(* Logix 5000 project; controller MV vendor 1 type 14 code 217 rev 31.11; software revision 31.00 *) (continued)
        [2].5   // Channel 1 extend button available
        [32].5   // CH1 run return flow check timer
        [26]   // CH1 no.of tank to be cleaned
        [31].0   // CH1 scavenge initialised
        [31].1   // CH1 prerinse initialised
        [32].4   // CH1 run return pump flag
        [34]   // CH1 command processor current step
        [38]   // CH1 pointer to DT service data file
        [11]   // CH1 route no.
        [33].2   // CH1 detergent tank high level probe covered
        [35]   // CH1 restart step
   MC_N100_20_alarm : ALARM_DIGITAL;
   MC_N100_20_Alarm_Ready : BOOL;
   MC_N100_20_Delayed_Timer2 : TIMER := (PRE := 1000);
   MC_N100_20_Fault_Returned : STRING;
   MC_N100_20_SQL_Done : DINT := -1;
   MC_N100_23_alarm : ALARM_DIGITAL;
   MC_N100_23_Alarm_Ready : BOOL;
   MC_N100_23_Delayed_Timer2 : TIMER := (PRE := 1000);
   MC_N100_23_Event_Returned : STRING := 'CH1_R1 feedbacks have failed.';
   MC_N100_23_Fault_Returned : STRING;
   MC_N100_23_SQL_Done : DINT := -1;
   MC_N100_29_0_Storagebit : BOOL;
   MC_N100_29_1_Storagebit : BOOL;
   MC_N100_29_2_Storagebit : BOOL;
   MC_N100_29_3_Storagebit : BOOL;
   MC_N100_29_4_Storagebit : BOOL;
   MC_N101 : INT[255];   // CH1 PC>PLC Channel 1 PC to PLC
        [0]   // CH1 PC button selected
        [0].2   // Stop channel 1 CIP selected
        [0].5   // Extend Channel 1 CIP selected
        [0].6   // Channel 1 end extend selected
        [0].15   // CH1 startup cancelled
        [0].7   // Channel 1 skip selected
        [0].4   // Abort channel 1 CIP selected
        [0].3   // Continue channel 1 CIP selected
        [0].1   // Start CH1 selected
        [0].0   // Initiate CH1 startup
   MC_N102 : INT[255] := ([1] := 1, [2] := 70, [3] := 1, [4] := 900, [5] := 1, [6] := 300, [10] := 2000, [11] := 90, [12] := 120, [13] := 7, [14] := 1, [15] := 6, [16] := 17, [17] := 1017, [19] := 11068, [21] := -1, [22] := -32768, [23] := -32768, [24] := -32768, [25] := -32768, [26] := -32768, [27] := -32768, [28] := -32768, [29] := -32768, [30] := -32768, [31] := -32768);   // CH1 PROG Channel 1 CIP progra m
        [1]   // CH1 no.prerinse cycles
        [10]   // CH1 CIP program flowrate setpoint (??/??)
        [14]   // CH1 CIP program detergent tank to use (1-2)
        [13].1   // CH1 recover rinse water flag
        [13].2   // CH1 use recovered water flag
        [0]   // CH1 scavenge time
        [15]   // CH1 CIP program route no.(1-6)
        [9]   // CH1 CIP program pressure setpoint (PSI)
        [16]   // CH1 CIP program program no.(1-47)
        [13].0   // CH1 Is Line Clean flag
        [21]   // CH1 CIP program vessel no.
        [4]   // CH1 detergent cycle time
        [6]   // CH1 postrinse cycle time
        [2]   // CH1 prerinse cycle time
        [3]   // CH1 no.detergent cycles
        [5]   // CH1 no.postrinse cycles
   MC_N103 : INT[255] := ([1] := 1, [2] := 2, [3] := 3, [4] := 4, [5] := 5, [6] := 6, [7] := 7, [8] := 8, [9] := 9, [10] := 10, [11] := 11, [12] := 12, [13] := 13, [14] := 14, [15] := 15, [16] := 16, [17] := 17, [18] := 18, [19] := 19, [20] := 64, [21] := 9999, [22] := 9999, [23] := 9999, [24] := 62, [25] := 99, [26] := -32768, [27] := 9999, [28] := 9999, [29] := 9999, [30] := 9999, [31] := -32768);   // CH1 ITEMS Chwd.nos.of items to be checked for Chan nel 1
        [0]   // CH1/R1 checkword no.
        [1]   // CH1/R2 checkword no.
        [2]   // CH1/R3 checkword no.
        [3]   // CH1/R4 checkword no.
        [4]   // CH1/R5 checkword no.
        [5]   // CH1/R6 checkword no.
        [12]   // CH1/DRAIN checkword no.
        [13]   // CH1/RR checkword no.
        [6]   // CH1/R1R checkword no.
        [7]   // CH1/R2R checkword no.
        [8]   // CH1/R3R checkword no.
        [9]   // CH1/R4R checkword no.
        [10]   // CH1/R5R checkword no.
        [11]   // CH1/R6R checkword no.
        [14]   // CH1/DR1 checkword no.
        [15]   // CH1/DR2 checkword no.
        [16]   // CH1/DT1 checkword no.
        [17]   // CH1/DT2 checkword no.
        [18]   // CH1/PR1 checkword no.
        [19]   // CH1/LF1 checkword no.
        [20]   // P1 checkword no.
   MC_N104 : INT[255] := ([0] := 6, [1] := 1017, [3] := 11068, [5] := 3, [6] := 14, [9] := 1);   // CH1 REPORT Channel 1 CIP report file
        [0].3   // CH1 final detergent strength save required
        [9]   // CH1 report detergent tank used (1 or 2)
        [0].0   // CH1 PLC -> PC save CIP report flag
        [0].1   // CH1 report save starting detergent strength flag
        [0].2   // CH1 report save final detergent strength flag
        [0]   // CH1 report flags
   MC_N108 : INT[255] := ([0] := 20, [1] := 8, [2] := 20, [3] := 4, [4] := 1);   // CH1 VDATA Channel 1 CIP progra m validation data
        [3]   // CH1 program validation loops this scan
        [4].0   // CH1 program validation complete flag
        [2]   // CH1 program validation loop counter
        [1]   // CH1 program validation max.loops per scan
        [4].1   // CH1 CIP program invalid flag
        [0]   // CH1 program validation CIP program size
        [4]   // CH1 program validation flags
   MC_N112 : INT[255] := ([0] := 1, [1] := 16, [2] := 3, [3] := -1, [4] := 2000, [9] := 5, [10] := 4, [11] := 16, [12] := 3, [13] := -1, [14] := -4, [40] := 4309, [42] := 20, [43] := 14, [44] := 137, [45] := 100, [48] := 23, [54] := 14641, [55] := 11826, [56] := 13873, [57] := 11832, [58] := 12338, [59] := 13102, [60] := 53, [101] := 6, [102] := 17, [103] := -1, [104] := 32);   // FVR DATA Data read from FV ro uting PLC
        [13]   // FV Routing CH2 fault register
        [4].0   // FV Routing > MV/FV CIP CH1 remote route open flag
        [102]   // CH1 current CIP program no.> Routing PLC
        [104].1   // CH1 CIP running flag > FV Routing PLC
        [104].4   // CH1 reset fault flag > FV Routing PLC
        [112]   // CH2 current CIP program no.> Routing PLC
        [114].1   // CH2 CIP running flag > FV Routing PLC
        [114].4   // CH2 reset fault flag > FV Routing PLC
        [104].3   // CH1 CIP complete flag > FV Routing PLC
        [114].3   // CH2 CIP complete flag > FV Routing PLC
        [103]   // CH1 no.of vessel being cleaned > Routing PLC
        [113]   // CH2 no.of vessel being cleaned > Routing PLC
        [4].1   // FV Routing > MV/FV CIP CH1 system reset flag
        [20].0   // Comms.to FV Routing PLC have failed
        [3]   // FV Routing CH1 fault register
        [0].0   // FV Routing > MV/FV CIP heartbeat
        [100].0   // MV/FV CIP > FV Routing heartbeat
        [104].0   // CH1 active flag > FV Routing PLC
        [104].6   // CH1 timing flag > FV Routing PLC
        [114].0   // CH2 active flag > FV Routing PLC
        [114].6   // CH2 timing flag > FV Routing PLC
        [14].1   // FV Routing > MV/FV CIP CH2 system reset flag
        [104].5   // CH1 detergent circulating flag > FV Routing PLC
        [114].5   // CH2 detergent circulating flag > FV Routing PLC
        [14].0   // FV Routing > MV/FV CIP CH2 remote route open flag
        [101]   // CH1 route no.> Routing PLC
        [104].2   // CH1 run return pump flag > FV Routing PLC
        [111]   // CH2 route no.> Routing PLC
        [114].2   // CH2 run return pump flag > FV Routing PLC
   MC_N113 : INT[255] := ([0] := 1, [1] := 1472, [2] := 511, [3] := -1, [11] := 1472, [12] := 511, [13] := -1, [40] := 4312, [42] := 20, [43] := 14, [44] := 137, [45] := 100, [48] := 23, [54] := 14641, [55] := 11826, [56] := 13873, [57] := 11832, [58] := 12338, [59] := 13102, [60] := 52, [101] := 6, [102] := 17, [103] := -1, [104] := 160);   // MVR DATA Data read from MV ro uting PLC
        [13]   // MV Routing CH2 fault register
        [4].0   // MV Routing > MV/FV CIP CH1 remote route open flag
        [104].1   // CH1 CIP running flag > FV Routing PLC
        [104].4   // CH1 reset fault flag > MV Routing PLC
        [114].1   // CH2 CIP running flag > MV Routing PLC
        [114].4   // CH2 reset fault flag > MV Routing PLC
        [104].3   // CH1 CIP complete flag > MV Routing PLC
        [114].3   // CH2 CIP complete flag > MV Routing PLC
        [4].1   // MV Routing > MV/FV CIP CH1 system reset flag
        [20].0   // Comms.to MV Routing PLC have failed
        [3]   // MV Routing CH1 fault register
        [0].0   // MV Routing > MV/FV CIP heartbeat
        [100].0   // MV/FV CIP > MV Routing heartbeat
        [104].0   // CH1 active flag > MV Routing PLC
        [104].5   // CH1 detergent circulating flag > MV Routing PLC
        [114].5   // CH2 detergent circulating flag > MV Routing PLC
        [14].0   // MV Routing > MV/FV CIP CH2 remote route open flag
        [114].0   // CH2 active flag > MV Routing PLC
        [14].1   // MV Routing > MV/FV CIP CH2 system reset flag
        [104].2   // CH1 run return pump flag > MV Routing PLC
        [114].2   // CH2 run return pump flag > MV Routing PLC
   MC_N114 : INT[255] := ([0] := 1, [20] := 1, [40] := -16384, [42] := 20, [43] := 14, [44] := 137, [45] := 100, [48] := 23, [54] := 14641, [55] := 11826, [56] := 13873, [57] := 11832, [58] := 12338, [59] := 13102, [60] := 56, [101] := 6, [102] := 17, [103] := -1, [104] := 32);   // YP DATA
        [104].1   // CH1 CIP running flag > Yeast Press PLC
        [104].4   // CH1 reset fault flag > Yeast Press PLC
        [14].1   // Yeast Press > MV/FV CIP CH2 system reset flag
        [114].1   // CH2 CIP running flag > Yeast Press PLC
        [114].4   // CH2 reset fault flag > Yeast Press PLC
        [104].5   // CH1 detergent circulating flag > Yeast Press PLC
        [114].5   // CH2 detergent circulating flag > Yeast Press PLC
        [4].0   // Yeast Press > MV/FV CIP CH1 remote route open flag
        [104].3   // CH1 CIP complete flag > Yeast Press PLC
        [100].0   // MV/FV CIP > Yeast Press heartbeat
        [104].0   // CH1 active flag > Yeast Press PLC
        [114].0   // CH2 active flag > Yeast Press PLC
        [114].3   // CH2 CIP complete flag > Yeast Press PLC
        [104].2   // CH1 run return pump flag > Yeast Press PLC
        [20].0   // Comms.to Yeast Press PLC have failed
        [13]   // Yeast Press CH2 fault register
        [114].2   // CH2 run return pump flag > Yeast Press PLC
        [4].1   // Yeast Press > MV/FV CIP CH1 system reset flag
        [0].0   // Yeast Press > MV/FV CIP heartbeat
        [3]   // Yeast Press CH1 fault register
   MC_N12 : INT[255];   // SYS_PARMS
        [28]   // PC>PLC Settings Current Day
        [0].0   // PLC>PC Settings Reload Request
        [27]   // PC>PLC Settings Current Month
        [32]   // Deferred chilling on fermentation delay (hrs.x10)
        [34]   // Deferred chilling on conditioning delay (hrs.x10)
        [1]   // PC>PLC settings Daily Rouse Start Hour
        [3]   // PC>PLC settings Daily Rouse Duration
        [2]   // PC>PLC settings Daily Rouse Start Minute
        [4]   // PC>PLC settings Hourly Rouse Duration
        [30]   // PC>PLC settings Current Minute
        [37]   // Deferred chilling off time hour
        [40]   // Deferred chilling maturation temp.high value
        [31]   // PC>PLC settings Current Second
        [38]   // Deferred chilling off time min.
        [33]   // Deferred chilling on maturation delay (hrs.x10)
        [35]   // Deferred chilling on time hour
        [36]   // Deferred chilling on time min.
        [26]   // PC>PLC Settings Current Year
        [29]   // PC>PLC settings Current Hour
        [39]   // Deferred chilling fermentation temp. high value
        [41]   // Deferred chilling conditioning temp. high value
   MC_N120 : INT[255] := ([0] := 1, [2] := 1, [20] := -1, [21] := 2, [22] := 2, [24] := 2, [25] := 2, [29] := 10, [38] := 90, [39] := 201);   // C2 PLC Channel 2 PLC data
        [31].2   // CH2 detergent initialised
        [31].3   // CH2 postrinse initialised
        [18].2   // CH2 return postrinse to detergent tank
        [32].2   // CH2 enable return pump off delay timer
        [0]   // CH2 status 0: Unavailable; 1: Idle; 2: Running; 3: Stopped; 4: Faulted
        [18].3   // CH2 enable postrinse return to detergent tank
        [32].8   // CH2 route return to detergent tank flag
        [18].0   // CH2 return flow on debounce timer
        [2].3   // Channel 2 continue button available
        [30].3   // CH2 run current cycle timer
        [18].1   // CH2 Is Detergent Return flag
        [2].6   // Channel 2 end extend available
        [6]   // CH2 current CIP total time minutes
        [7]   // CH2 current CIP total time seconds
        [10]   // CH2 detergent tank to use (1 or 2)
        [32].9   // CH2 initialise supply pump PID flag
        [28].0   // CH2 MV Routing PLC in use flag
        [28].1   // CH2 FV Routing PLC in use flag
        [12]   // CH2 current CIP program no.
        [2].0   // Channel 2 start button available
        [30].4   // CH2 cycle complete flag
        [27].3   // CH2 drive new route 3 routing valves
        [27].4   // CH2 drive new route 4 routing valves
        [27].5   // CH2 drive new route 5 routing valves
        [27].6   // CH2 drive new route 6 routing valves
        [19].1   // P2 PID pressure control selected
        [19].3   // P2 PID flowrate control selected
        [33].4   // CH2 detergent tank low level probe uncovered
        [32].6   // CH2 run detergent return check timer
        [33].0   // CH2 open detergent tank return valve
        [33].1   // CH2 open detergent tank outlet valve
        [2].1   // CH2 startup in progress
        [30].2   // Channel 2 initialised
        [30].5   // CH2 extend cycle flag
        [31].10   // CH2 detergent active
        [31].11   // CH2 postrinse active
        [32].3   // CH2 open supply route flag
        [20]   // CH2 fault register
        [23]   // CH2 event register
        [32].7   // CH2 open return route flag
        [30].0   // CH2 reset flag
        [32].1   // CH2 enable return pump on delay timer
        [8]   // CH2 current CIP total stopped time minutes
        [9]   // CH2 current CIP total stopped time seconds
        [4]   // CH2 total subcycles to do
        [17]   // CH2 current substep
        [19]   // CH2 PID flags /0: Press.inhibited /1: Press.selected /2: Flow inhibited /3: Flow selected
        [2].2   // Channel 2 stop button available
        [30].1   // CH2 active flag
        [2].4   // Channel 2 abort button availble
        [2].7   // Channel 2 skip button available
        [33].3   // CH2 detergent tank working level probe covered
        [1]   // CH2 current CIP cycle
        [21]   // CH2 fault parameter #1
        [22]   // CH2 fault parameter #2
        [24]   // CH2 event parameter #1
        [31].8   // CH2 scavenge active
        [18].4   // CH2 waiting for DT service flag
        [33].2   // CH2 detergent tank high level probe covered
        [28].2   // CH2 Yeast Press PLC in use flag
        [2].5   // Channel 2 extend button available
        [32].5   // CH2 run return flow check timer
        [31].9   // CH2 prerinse active
        [26]   // CH2 no.of tank to be cleaned
        [3]   // CH2 current subcycle no.
        [5]   // CH2 time left this cycle
        [31].0   // CH2 scavenge initialised
        [34]   // CH2 command processor current step
        [38]   // CH2 pointer to DT service data file
        [31].1   // CH2 prerinse initialised
        [32].4   // CH2 run return pump flag
        [11]   // CH2 route no.
        [35]   // CH2 restart step
   MC_N120_20_alarm : ALARM_DIGITAL;
   MC_N120_20_Alarm_Ready : BOOL;
   MC_N120_20_Delayed_Timer2 : TIMER := (PRE := 1000);
   MC_N120_20_Fault_Returned : STRING;
   MC_N120_20_SQL_Done : DINT := -1;
   MC_N120_23_alarm : ALARM_DIGITAL;
   MC_N120_23_Alarm_Ready : BOOL;
   MC_N120_23_Delayed_Timer2 : TIMER := (PRE := 1000);
   MC_N120_23_Event_Returned : STRING := 'CH1_R1 feedbacks have failed.';
   MC_N120_23_SQL_Done : DINT := -1;
   MC_N120_29_0_Storagebit : BOOL;
   MC_N120_29_1_Storagebit : BOOL;
   MC_N120_29_2_Storagebit : BOOL;
   MC_N120_29_3_Storagebit : BOOL;
   MC_N120_29_4_Storagebit : BOOL;
   MC_N121 : INT[255];   // CH2 PC>PLC Channel 2 PC to PLC
        [0]   // CH2 PC button selected
        [0].2   // Stop channel 2 CIP selected
        [0].5   // Extend Channel 2 CIP selected
        [0].6   // Channel 2 end extend selected
        [0].15   // CH2 startup cancelled
        [0].7   // Channel 2 skip selected
        [0].4   // Abort channel 2 CIP selected
        [0].3   // Continue channel 2 CIP selected
        [0].1   // Start CH2 selected
        [0].0   // Initiate CH2 startup
   MC_N122 : INT[255] := ([0] := -32768, [1] := -32768, [2] := -32768, [3] := -32768, [4] := -32768, [5] := -32768, [6] := -32768, [7] := -32768, [8] := -32768, [9] := -32768, [10] := -32768, [11] := -32768, [12] := -32768, [13] := -32768, [14] := -32768, [15] := -32768, [16] := -32768, [17] := -32768, [18] := -32768, [19] := -32768, [20] := -32768, [21] := -32768, [22] := -32768, [23] := -32768, [24] := -32768, [25] := -32768, [26] := -32768, [27] := -32768, [28] := -32768, [29] := -32768, [30] := -32768, [31] := -32768);   // CH2 PROG Channel 2 CIP progra m
        [1]   // CH2 no.prerinse cycles
        [10]   // CH2 CIP program flowrate setpoint (??/??)
        [14]   // CH2 CIP program detergent tank to use (1-2)
        [13].1   // CH2 recover rinse water flag
        [13].2   // CH2 use recovered water flag
        [15]   // CH2 CIP program route no.(1-6)
        [0]   // CH2 scavenge time
        [9]   // CH2 CIP program pressure setpoint (PSI)
        [16]   // CH2 CIP program program no.(1-47)
        [4]   // CH2 detergent cycle time
        [6]   // CH2 postrinse cycle time
        [13].0   // CH2 Is Line Clean flag
        [21]   // CH2 CIP program vessel no.
        [2]   // CH2 prerinse cycle time
        [3]   // CH2 no.detergent cycles
        [5]   // CH2 no.postrinse cycles
   MC_N123 : INT[255] := ([0] := 20, [1] := 21, [2] := 22, [3] := 23, [4] := 24, [5] := 25, [6] := 26, [7] := 27, [8] := 28, [9] := 29, [10] := 30, [11] := 31, [12] := 32, [13] := 33, [14] := 34, [15] := 35, [16] := 36, [17] := 37, [18] := 38, [19] := 39, [20] := 65, [21] := 9999, [22] := 9999, [23] := 9999, [24] := 68, [25] := 81, [26] := -32768, [27] := 9999, [28] := 9999, [29] := 9999, [30] := 9999, [31] := -32768);   // CH2 ITEMS Chwd.nos.of items to be checked for Chan nel 2
        [0]   // CH2/R1 checkword no.
        [1]   // CH2/R2 checkword no.
        [2]   // CH2/R3 checkword no.
        [3]   // CH2/R4 checkword no.
        [4]   // CH2/R5 checkword no.
        [5]   // CH2/R6 checkword no.
        [12]   // CH2/DRAIN checkword no.
        [13]   // CH2/RR checkword no.
        [6]   // CH2/R1R checkword no.
        [7]   // CH2/R2R checkword no.
        [8]   // CH2/R3R checkword no.
        [9]   // CH2/R4R checkword no.
        [10]   // CH2/R5R checkword no.
        [11]   // CH2/R6R checkword no.
        [14]   // CH2/DR1 checkword no.
        [15]   // CH2/DR2 checkword no.
        [16]   // CH2/DT1 checkword no.
        [17]   // CH2/DT2 checkword no.
        [18]   // CH2/PR1 checkword no.
        [19]   // CH2/LF1 checkword no.
        [20]   // P2 checkword no.
   MC_N124 : INT[255] := ([0] := 14, [1] := 15, [3] := 11065, [5] := 20, [6] := 45, [9] := 2);   // CH2 REPORT Channel 2 CIP report file
        [0].0   // CH2 PLC -> PC save CIP report flag
        [0].3   // CH2 final detergent strength save required
        [9]   // CH2 report detergent tank used (1 or 2)
        [0].1   // CH2 report save starting detergent strength flag
        [0].2   // CH2 report save final detergent strength flag
        [0]   // CH2 report flags
   MC_N128 : INT[255] := ([0] := 20, [1] := 8, [2] := 20, [3] := 4, [4] := 1);   // CH2 VDATA Channel 2 CIP progra m validation data
        [3]   // CH2 program validation loops this scan
        [2]   // CH2 program validation loop counter
        [4].0   // CH2 program validation complete flag
        [1]   // CH2 program validation max.loops per scan
        [4].1   // CH2 CIP program invalid flag
        [0]   // CH2 program validation CIP program size
        [4]   // CH2 program validation flags
   MC_N140 : INT[31] := ([0] := 1, [1] := 1, [23] := -1, [24] := -1, [25] := 30);   // RT FILL RT filling routine d ata
        [12]   // RT/FTX01 volume count (hl.x 10)
        [16]   // RT filling max.flush volume
        [1].1   // RT filling startup in progress
        [6].1   // RT filling source vessel is CT
        [7]   // RT filling destination vessel no.
        [20]   // GEA vessel pointer
        [1].3   // RT filling Continue button available
        [6].4   // RT filling source is GEA MV
        [6].5   // RT filling source is GEA CT
        [6].0   // RT filling source vessel is old MV
        [1].12   // RT filling extend transfer available
        [5]   // RT filling command processor current step
        [1].10   // Enable Water Flush button available
        [1].11   // Disable MV Water Flush button available
        [1].8   // RT filling End Transfer button available
        [4].7   // RT filling beer/ liquor changeover flag
        [1].5   // RTfilling Confirm RT Vent Valve Open button available
        [18]   // Finings total dosed for PC display (ltr.x 10)
        [1].14   // RT filling audible alarm off button available
        [4].10   // RT filling destination RT high volume reached
        [6].2   // RT filling source vessel is new MV
        [15]   // RT filling pointer to destination RT's data file
        [1].6   // RT filling Confirm Liquor Flush Initiated button available
        [1].2   // RT filling Stop button available
        [14]   // RT filling max. transfer volume
        [4].6   // RT filling open route to RT flag
        [4].9   // RT filling destination vessel high level
        [1].0   // RT filling Start button available
        [6].3   // RT filling filling via filter flag
        [4].8   // Beer at CTX probe RT/CTX01
        [1].13   // RT filling flush available
        [9]   // RT filling MV packing line no.
        [17]   // RT filling finings volume error (pts.x10/brl.)
        [1].7   // Confirm Transfer Complete button available
        [4].11   // RT filling destination RT high level alarm
        [4].14   // RT filling ignore new MV tank empty flag
        [4].12   // RT filling Drive MV Water Flush Valve flag
        [4].13   // RT filling drive audible alarm/ beacon flag
        [1].9   // RT filling Select New Destination RT button available
        [1].4   // RT filling Abort button available
        [23]   // RT filling fault register
        [13]   // RT filling route volume
        [4].0   // RT filling reset flag
        [24]   // RT filling event register
        [10]   // RT filling transfer volume
        [25]   // RT filling work register
        [4].1   // RT filling active flag
        [4].2   // RT filling initialised
        [8]   // RT filling source vessel no.
        [2]   // RT filling current step
        [3]   // RT filling restart step
        [0]   // RT filling status 0: Unavailable; 1: Idle; 2: Running; 3: Stopped; 4: Fault 5: Waiting
   MC_N160 : INT[255] := ([0] := -32768, [1] := 9999, [2] := 9999, [3] := 9999, [4] := 9999, [5] := 9999, [6] := 9999, [7] := -32768);   // P40 CHECK
   MC_N161 : INT[255] := ([0] := -32768, [1] := 9999, [2] := 9999, [3] := 9999, [4] := 9999, [5] := 9999, [6] := 9999, [7] := -32768);   // P41 CHECK
   MC_N162 : INT[255] := ([0] := 63, [1] := -32768, [2] := 9999, [3] := 9999, [4] := 9999, [5] := 9999, [6] := 9999, [7] := -32768);   // P42 CHECK
   MC_N163 : INT[255] := ([0] := -32768, [1] := 9999, [2] := 9999, [3] := 9999, [4] := 9999, [5] := 9999, [6] := 9999, [7] := -32768);   // P43 CHECK
   MC_N164 : INT[255] := ([0] := -32768, [1] := 9999, [2] := 9999, [3] := 9999, [4] := 9999, [5] := 9999, [6] := 9999, [7] := -32768);   // P44 CHECK
   MC_N165 : INT[255] := ([0] := -32768, [1] := 9999, [2] := 9999, [3] := 9999, [4] := 9999, [5] := 9999, [6] := 9999, [7] := -32768);   // P45 CHECK
   MC_N166 : INT[255] := ([0] := -32768, [1] := 9999, [2] := 9999, [3] := 9999, [4] := 9999, [5] := 9999, [6] := 9999, [7] := -32768);   // P46 CHECK
   MC_N167 : INT[255] := ([0] := -32768, [1] := 9999, [2] := 9999, [3] := 9999, [4] := 9999, [5] := 9999, [6] := 9999, [7] := -32768);   // Original N File From SLC, No Description Available
   MC_N20 : INT[255] := ([0] := 1531, [1] := -32765, [2] := 650, [3] := 10, [8] := 1500, [12] := 100, [14] := 558, [15] := 92, [18] := -3898, [19] := -3372, [21] := 7520, [22] := 5040, [25] := 1638, [27] := 650, [28] := 400, [31] := 3, [32] := 3, [34] := 9150, [36] := 92);   // P1 PRESS Control block and da ta for P1 pressure P ID loop
        [37]   // P1 pressure PID saved op.mode
        [31].1   // P1 pressure PID loop high absolute alarm flag
        [31].0   // P1 pressure PID loop deviation alarm flag
        [30]   // P1 pressure PID loop deviation alarm setting
        [26]   // P1 pressure PID loop PLC output
        [38]   // P1 pressure PID saved PLC output
        [25]   // P1 pressure PID loop local (PC) output
        [2]   // P1 pressure PID loop setpoint
        [0].1   // P1 pressure PID loop auto/manual flag
        [28]   // P1 pressure PID loop high absolute alarm setting
        [31].2   // P1 pressure PID loop low absolute alarm flag
        [14]   // P1 pressure PID loop process variable
        [23]   // P1 press.op.mode: 0: PLC manual; 1: PLC setpoint; 2: Local manual; 3: Local setpoint;
        [24]   // P1 pressure PID loop local (PC) setpoint
        [27]   // P1 pressure PID loop PLC setpoint
        [35]   // P1 pressure PID loop desired output
        [29]   // P1 pressure PID loop low absolute alarm setting
        [36]   // Work register
   MC_N200 : INT[255] := ([0] := 103, [1] := -1, [2] := 26, [3] := 99);   // CHK_WORK Plant item fault che cking work area
        [0]   // Item checking routine file pointer
        [1]   // Faulted plant item checkword no.
   MC_N201 : INT[255] := ([0] := 68, [1] := 81, [2] := -32768, [3] := 9999, [4] := 9999, [5] := 9999, [6] := 9999, [7] := -32768);   // P1 CHECK CIP program 1 plant item check list
   MC_N202 : INT[255] := ([0] := 71, [1] := 61, [2] := 98, [3] := -32768, [4] := 9999, [5] := 9999, [6] := 9999, [7] := -32768);   // P2 CHECK CIP program 2 plant item check list
   MC_N203 : INT[255] := ([0] := 72, [1] := 61, [2] := 98, [3] := -32768, [4] := 9999, [5] := 9999, [6] := 9999, [7] := -32768);   // P3 CHECK CIP program 3 plant item check list
   MC_N204 : INT[255] := ([0] := 69, [1] := -32768, [2] := 9999, [3] := 9999, [4] := 9999, [5] := 9999, [6] := 9999, [7] := -32768);   // P4 CHECK CIP program 4 plant item check list
   MC_N205 : INT[255] := ([0] := 69, [1] := -32768, [2] := 9999, [3] := 9999, [4] := 9999, [5] := 9999, [6] := 9999, [7] := -32768);   // P5 CHECK CIP program 5 plant item check list
   MC_N206 : INT[255] := ([0] := 69, [1] := -32768, [2] := 9999, [3] := 9999, [4] := 9999, [5] := 9999, [6] := 9999, [7] := -32768);   // P6 CHECK CIP program 6 plant item check list
   MC_N207 : INT[255] := ([0] := -32768, [1] := 9999, [2] := 9999, [3] := 9999, [4] := 9999, [5] := 9999, [6] := 9999, [7] := -32768);   // P7 CHECK CIP program 7 plant item check list
   MC_N208 : INT[255] := ([0] := 59, [1] := 96, [2] := -32768, [3] := 9999, [4] := 9999, [5] := 9999, [6] := 9999, [7] := -32768);   // P8 CHECK CIP program 8 plant item check list
   MC_N209 : INT[255] := ([0] := 59, [1] := 96, [2] := -32768, [3] := 9999, [4] := 9999, [5] := 9999, [6] := 9999, [7] := -32768);   // P9 CHECK CIP program 9 plant item check list
   MC_N21 : INT[255] := ([1] := -31733, [2] := 2000, [3] := 5, [8] := 5000, [11] := 100, [12] := 10, [13] := 20, [14] := 1995, [15] := 5, [16] := 72, [17] := -4096, [18] := 25212, [21] := 5041, [22] := 3500, [23] := 1, [24] := 5000, [25] := 12287, [27] := 2000, [31] := 3, [34] := 6538, [35] := 11832, [36] := 5, [37] := 1);   // P1 FLOW Control block and da ta for P1 flowrate P ID loop
        [37]   // P1 flowrate PID saved op.mode
        [31].1   // P1 flowrate PID loop high absolute alarm flag
        [31].0   // P1 flowrate PID loop deviation alarm flag
        [30]   // P1 flowrate PID loop deviation alarm setting
        [28]   // P1 flowrate PID loop high absolute alarm setting
        [38]   // P1 flowrate PID saved PLC output
        [26]   // P1 flowrate PID loop PLC output
        [14]   // P1 flowrate PID loop process variable
        [25]   // P1 flowrate PID loop local (PC) output
        [2]   // P1 flowrate PID loop setpoint
        [0].1   // P1 flowrate PID loop auto/manual flag
        [31].2   // P1 flowrate PID loop low absolute alarm flag
        [24]   // P1 flowrate PID loop local (PC) setpoint
        [27]   // P1 flowrate PID loop PLC setpoint
        [29]   // P1 flowrate PID loop low absolute alarm setting
        [35]   // P1 flowrate PID loop desired output
        [23]   // P1 flow op.mode: 0: PLC manual; 1: PLC setpoint; 2: Local manual; 3: Local setpoint;
        [36]   // Work register
   MC_N210 : INT[255] := ([0] := 60, [1] := 97, [2] := -32768, [3] := 9999, [4] := 9999, [5] := 9999, [6] := 9999, [7] := -32768);   // P10 CHECK CIP program 10 plant item check list
   MC_N211 : INT[255] := ([0] := 60, [1] := 97, [2] := -32768, [3] := 9999, [4] := 9999, [5] := 9999, [6] := 9999, [7] := -32768);   // P11 CHECK CIP program 11 plant item check list
   MC_N212 : INT[255] := ([0] := 73, [1] := 47, [2] := 62, [3] := 99, [4] := -32768, [5] := 9999, [6] := 9999, [7] := -32768);   // P12 CHECK CIP program 12 plant item check list
   MC_N213 : INT[255] := ([0] := 74, [1] := 48, [2] := 62, [3] := 99, [4] := -32768, [5] := 9999, [6] := 9999, [7] := -32768);   // P13 CHECK CIP program 13 plant item check list
   MC_N214 : INT[255] := ([0] := 75, [1] := 49, [2] := 62, [3] := 99, [4] := -32768, [5] := 9999, [6] := 9999, [7] := -32768);   // P14 CHECK CIP program 14 plant item check list
   MC_N215 : INT[255] := ([0] := 76, [1] := 50, [2] := 62, [3] := 99, [4] := -32768, [5] := 9999, [6] := 9999, [7] := -32768);   // P15 CHECK CIP program 15 plant item check list
   MC_N216 : INT[255] := ([0] := 77, [1] := 51, [2] := 62, [3] := 99, [4] := -32768, [5] := 9999, [6] := 9999, [7] := -32768);   // P16 CHECK CIP program 16 plant item check list
   MC_N217 : INT[255] := ([0] := 62, [1] := 99, [2] := -32768, [3] := 9999, [4] := 9999, [5] := 9999, [6] := 9999, [7] := -32768);   // P17 CHECK CIP program 17 plant item check list
   MC_N218 : INT[255] := ([0] := 60, [1] := 97, [2] := -32768, [3] := 9999, [4] := 9999, [5] := 9999, [6] := 9999, [7] := -32768);   // P18 CHECK CIP program 18 plant item check list
   MC_N219 : INT[255] := ([0] := 59, [1] := 96, [2] := -32768, [3] := 9999, [4] := 9999, [5] := 9999, [6] := 9999, [7] := -32768);   // P19 CHECK CIP program 19 plant item check list
   MC_N22 : INT[255] := ([0] := -32765, [2] := 450, [3] := 1, [7] := 1500, [11] := 100, [13] := 20, [14] := 84, [15] := 366, [17] := -4820, [18] := -9972, [20] := 13744, [21] := 5041, [22] := 520, [24] := 600, [25] := 8192, [27] := 450, [30] := 50, [31] := 3, [34] := 1369, [36] := 366);   // P2 PRESS Control block and da ta for P2 pressure P ID loop
        [37]   // P2 pressure PID saved op.mode
        [31].1   // P2 pressure PID loop high absolute alarm flag
        [31].0   // P2 pressure PID loop deviation alarm flag
        [28]   // P2 pressure PID loop high absolute alarm setting
        [31].2   // P2 pressure PID loop low absolute alarm flag
        [30]   // P2 pressure PID loop deviation alarm setting
        [24]   // P2 pressure PID loop local (PC) setpoint
        [38]   // P2 pressure PID saved PLC output
        [26]   // P2 pressure PID loop PLC output
        [14]   // P2 pressure PID loop process variable
        [25]   // P2 pressure PID loop local (PC) output
        [2]   // P2 pressure PID loop setpoint
        [0].1   // P2 pressure PID loop auto/manual flag
        [27]   // P2 pressure PID loop PLC setpoint
        [23]   // P2 press.op.mode: 0: PLC manual; 1: PLC setpoint; 2: Local manual; 3: Local setpoint;
        [29]   // P2 pressure PID loop low absolute alarm setting
        [35]   // P2 pressure PID loop desired output
        [36]   // Work register
   MC_N220 : INT[255] := ([0] := 59, [1] := 96, [2] := -32768, [3] := 9999, [4] := 9999, [5] := 9999, [6] := 9999, [7] := -32768);   // P20 CHECK CIP program 20 plant item check list
   MC_N221 : INT[255] := ([0] := 59, [1] := 96, [2] := -32768, [3] := 9999, [4] := 9999, [5] := 9999, [6] := 9999, [7] := -32768);   // P21 CHECK CIP program 21 plant item check list
   MC_N222 : INT[255] := ([0] := 70, [1] := 59, [2] := 96, [3] := -32768, [4] := 9999, [5] := 9999, [6] := 9999, [7] := -32768);   // P22 CHECK CIP program 22 plant item check list
   MC_N223 : INT[255] := ([0] := 70, [1] := 59, [2] := 96, [3] := -32768, [4] := 9999, [5] := 9999, [6] := 9999, [7] := -32768);   // P23 CHECK CIP program 23 plant item check list
